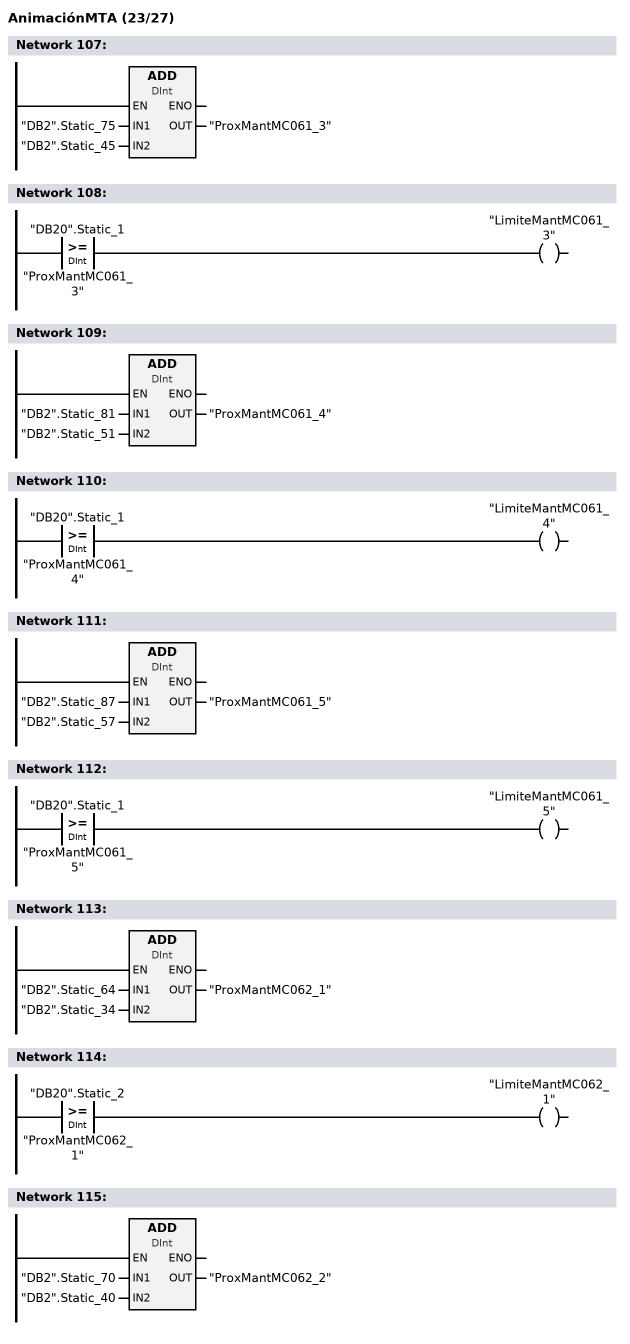
   RUNG wire#powerrail
      { S7_Templates := "SrcType := DInt"; S7_GenerateENO := "TRUE" } Add(in1 := "DB2".Static_75, in2 := "DB2".Static_45, out => "ProxMantMC061_3")
   END_RUNG
   // the same network as SCL:
   "ProxMantMC061_3" := "DB2".Static_75 + "DB2".Static_45;
END_REGION

REGION Network 108
   RUNG wire#powerrail
      { S7_Templates := "SrcType := DInt" } GE_Contact(in1 := "DB20".Static_1, in2 := "ProxMantMC061_3")
      Coil( "LimiteMantMC061_3" )
   END_RUNG
   // the same network as SCL:
   "LimiteMantMC061_3" := "DB20".Static_1 >= "ProxMantMC061_3";
END_REGION

REGION Network 109
   RUNG wire#powerrail
      { S7_Templates := "SrcType := DInt"; S7_GenerateENO := "TRUE" } Add(in1 := "DB2".Static_81, in2 := "DB2".Static_51, out => "ProxMantMC061_4")
   END_RUNG
   // the same network as SCL:
   "ProxMantMC061_4" := "DB2".Static_81 + "DB2".Static_51;
END_REGION

REGION Network 110
   RUNG wire#powerrail
      { S7_Templates := "SrcType := DInt" } GE_Contact(in1 := "DB20".Static_1, in2 := "ProxMantMC061_4")
      Coil( "LimiteMantMC061_4" )
   END_RUNG
   // the same network as SCL:
   "LimiteMantMC061_4" := "DB20".Static_1 >= "ProxMantMC061_4";
END_REGION

REGION Network 111
   RUNG wire#powerrail
      { S7_Templates := "SrcType := DInt"; S7_GenerateENO := "TRUE" } Add(in1 := "DB2".Static_87, in2 := "DB2".Static_57, out => "ProxMantMC061_5")
   END_RUNG
   // the same network as SCL:
   "ProxMantMC061_5" := "DB2".Static_87 + "DB2".Static_57;
END_REGION

REGION Network 112
   RUNG wire#powerrail
      { S7_Templates := "SrcType := DInt" } GE_Contact(in1 := "DB20".Static_1, in2 := "ProxMantMC061_5")
      Coil( "LimiteMantMC061_5" )
   END_RUNG
   // the same network as SCL:
   "LimiteMantMC061_5" := "DB20".Static_1 >= "ProxMantMC061_5";
END_REGION

REGION Network 113
   RUNG wire#powerrail
      { S7_Templates := "SrcType := DInt"; S7_GenerateENO := "TRUE" } Add(in1 := "DB2".Static_64, in2 := "DB2".Static_34, out => "ProxMantMC062_1")
   END_RUNG
   // the same network as SCL:
   "ProxMantMC062_1" := "DB2".Static_64 + "DB2".Static_34;
END_REGION

REGION Network 114
   RUNG wire#powerrail
      { S7_Templates := "SrcType := DInt" } GE_Contact(in1 := "DB20".Static_2, in2 := "ProxMantMC062_1")
      Coil( "LimiteMantMC062_1" )
   END_RUNG
   // the same network as SCL:
   "LimiteMantMC062_1" := "DB20".Static_2 >= "ProxMantMC062_1";
END_REGION

REGION Network 115
   RUNG wire#powerrail
      { S7_Templates := "SrcType := DInt"; S7_GenerateENO := "TRUE" } Add(in1 := "DB2".Static_70, in2 := "DB2".Static_40, out => "ProxMantMC062_2")
   END_RUNG
   // the same network as SCL:
   "ProxMantMC062_2" := "DB2".Static_70 + "DB2".Static_40;
END_REGION

REGION Network 116
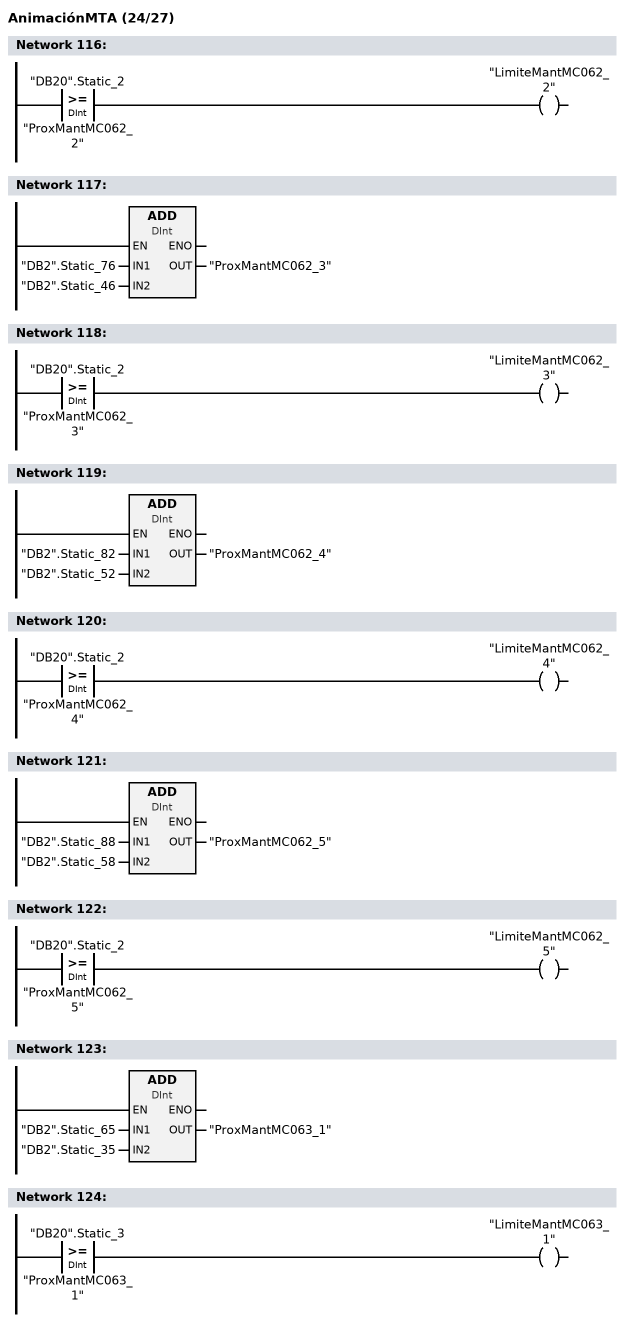
   RUNG wire#powerrail
      { S7_Templates := "SrcType := DInt" } GE_Contact(in1 := "DB20".Static_2, in2 := "ProxMantMC062_2")
      Coil( "LimiteMantMC062_2" )
   END_RUNG
   // the same network as SCL:
   "LimiteMantMC062_2" := "DB20".Static_2 >= "ProxMantMC062_2";
END_REGION

REGION Network 117
   RUNG wire#powerrail
      { S7_Templates := "SrcType := DInt"; S7_GenerateENO := "TRUE" } Add(in1 := "DB2".Static_76, in2 := "DB2".Static_46, out => "ProxMantMC062_3")
   END_RUNG
   // the same network as SCL:
   "ProxMantMC062_3" := "DB2".Static_76 + "DB2".Static_46;
END_REGION

REGION Network 118
   RUNG wire#powerrail
      { S7_Templates := "SrcType := DInt" } GE_Contact(in1 := "DB20".Static_2, in2 := "ProxMantMC062_3")
      Coil( "LimiteMantMC062_3" )
   END_RUNG
   // the same network as SCL:
   "LimiteMantMC062_3" := "DB20".Static_2 >= "ProxMantMC062_3";
END_REGION

REGION Network 119
   RUNG wire#powerrail
      { S7_Templates := "SrcType := DInt"; S7_GenerateENO := "TRUE" } Add(in1 := "DB2".Static_82, in2 := "DB2".Static_52, out => "ProxMantMC062_4")
   END_RUNG
   // the same network as SCL:
   "ProxMantMC062_4" := "DB2".Static_82 + "DB2".Static_52;
END_REGION

REGION Network 120
   RUNG wire#powerrail
      { S7_Templates := "SrcType := DInt" } GE_Contact(in1 := "DB20".Static_2, in2 := "ProxMantMC062_4")
      Coil( "LimiteMantMC062_4" )
   END_RUNG
   // the same network as SCL:
   "LimiteMantMC062_4" := "DB20".Static_2 >= "ProxMantMC062_4";
END_REGION

REGION Network 121
   RUNG wire#powerrail
      { S7_Templates := "SrcType := DInt"; S7_GenerateENO := "TRUE" } Add(in1 := "DB2".Static_88, in2 := "DB2".Static_58, out => "ProxMantMC062_5")
   END_RUNG
   // the same network as SCL:
   "ProxMantMC062_5" := "DB2".Static_88 + "DB2".Static_58;
END_REGION

REGION Network 122
   RUNG wire#powerrail
      { S7_Templates := "SrcType := DInt" } GE_Contact(in1 := "DB20".Static_2, in2 := "ProxMantMC062_5")
      Coil( "LimiteMantMC062_5" )
   END_RUNG
   // the same network as SCL:
   "LimiteMantMC062_5" := "DB20".Static_2 >= "ProxMantMC062_5";
END_REGION

REGION Network 123
   RUNG wire#powerrail
      { S7_Templates := "SrcType := DInt"; S7_GenerateENO := "TRUE" } Add(in1 := "DB2".Static_65, in2 := "DB2".Static_35, out => "ProxMantMC063_1")
   END_RUNG
   // the same network as SCL:
   "ProxMantMC063_1" := "DB2".Static_65 + "DB2".Static_35;
END_REGION

REGION Network 124
   RUNG wire#powerrail
      { S7_Templates := "SrcType := DInt" } GE_Contact(in1 := "DB20".Static_3, in2 := "ProxMantMC063_1")
      Coil( "LimiteMantMC063_1" )
   END_RUNG
   // the same network as SCL:
   "LimiteMantMC063_1" := "DB20".Static_3 >= "ProxMantMC063_1";
END_REGION

REGION Network 125
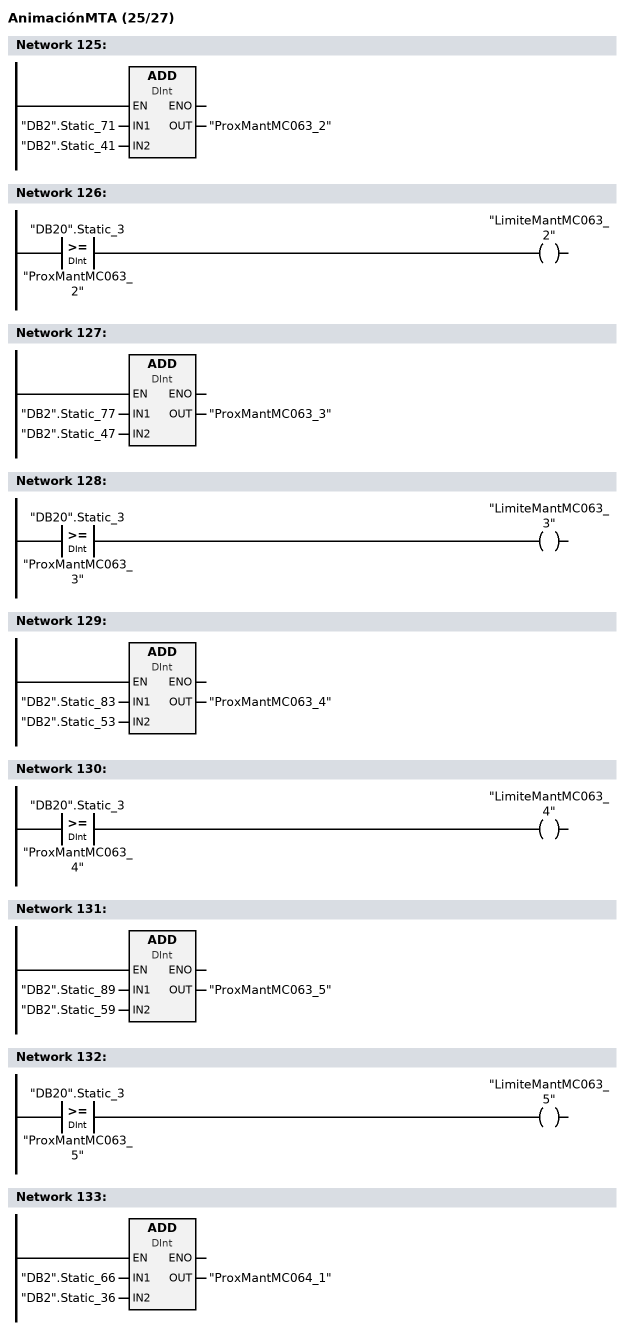
   RUNG wire#powerrail
      { S7_Templates := "SrcType := DInt"; S7_GenerateENO := "TRUE" } Add(in1 := "DB2".Static_71, in2 := "DB2".Static_41, out => "ProxMantMC063_2")
   END_RUNG
   // the same network as SCL:
   "ProxMantMC063_2" := "DB2".Static_71 + "DB2".Static_41;
END_REGION

REGION Network 126
   RUNG wire#powerrail
      { S7_Templates := "SrcType := DInt" } GE_Contact(in1 := "DB20".Static_3, in2 := "ProxMantMC063_2")
      Coil( "LimiteMantMC063_2" )
   END_RUNG
   // the same network as SCL:
   "LimiteMantMC063_2" := "DB20".Static_3 >= "ProxMantMC063_2";
END_REGION

REGION Network 127
   RUNG wire#powerrail
      { S7_Templates := "SrcType := DInt"; S7_GenerateENO := "TRUE" } Add(in1 := "DB2".Static_77, in2 := "DB2".Static_47, out => "ProxMantMC063_3")
   END_RUNG
   // the same network as SCL:
   "ProxMantMC063_3" := "DB2".Static_77 + "DB2".Static_47;
END_REGION

REGION Network 128
   RUNG wire#powerrail
      { S7_Templates := "SrcType := DInt" } GE_Contact(in1 := "DB20".Static_3, in2 := "ProxMantMC063_3")
      Coil( "LimiteMantMC063_3" )
   END_RUNG
   // the same network as SCL:
   "LimiteMantMC063_3" := "DB20".Static_3 >= "ProxMantMC063_3";
END_REGION

REGION Network 129
   RUNG wire#powerrail
      { S7_Templates := "SrcType := DInt"; S7_GenerateENO := "TRUE" } Add(in1 := "DB2".Static_83, in2 := "DB2".Static_53, out => "ProxMantMC063_4")
   END_RUNG
   // the same network as SCL:
   "ProxMantMC063_4" := "DB2".Static_83 + "DB2".Static_53;
END_REGION

REGION Network 130
   RUNG wire#powerrail
      { S7_Templates := "SrcType := DInt" } GE_Contact(in1 := "DB20".Static_3, in2 := "ProxMantMC063_4")
      Coil( "LimiteMantMC063_4" )
   END_RUNG
   // the same network as SCL:
   "LimiteMantMC063_4" := "DB20".Static_3 >= "ProxMantMC063_4";
END_REGION

REGION Network 131
   RUNG wire#powerrail
      { S7_Templates := "SrcType := DInt"; S7_GenerateENO := "TRUE" } Add(in1 := "DB2".Static_89, in2 := "DB2".Static_59, out => "ProxMantMC063_5")
   END_RUNG
   // the same network as SCL:
   "ProxMantMC063_5" := "DB2".Static_89 + "DB2".Static_59;
END_REGION

REGION Network 132
   RUNG wire#powerrail
      { S7_Templates := "SrcType := DInt" } GE_Contact(in1 := "DB20".Static_3, in2 := "ProxMantMC063_5")
      Coil( "LimiteMantMC063_5" )
   END_RUNG
   // the same network as SCL:
   "LimiteMantMC063_5" := "DB20".Static_3 >= "ProxMantMC063_5";
END_REGION

REGION Network 133
   RUNG wire#powerrail
      { S7_Templates := "SrcType := DInt"; S7_GenerateENO := "TRUE" } Add(in1 := "DB2".Static_66, in2 := "DB2".Static_36, out => "ProxMantMC064_1")
   END_RUNG
   // the same network as SCL:
   "ProxMantMC064_1" := "DB2".Static_66 + "DB2".Static_36;
END_REGION

REGION Network 134
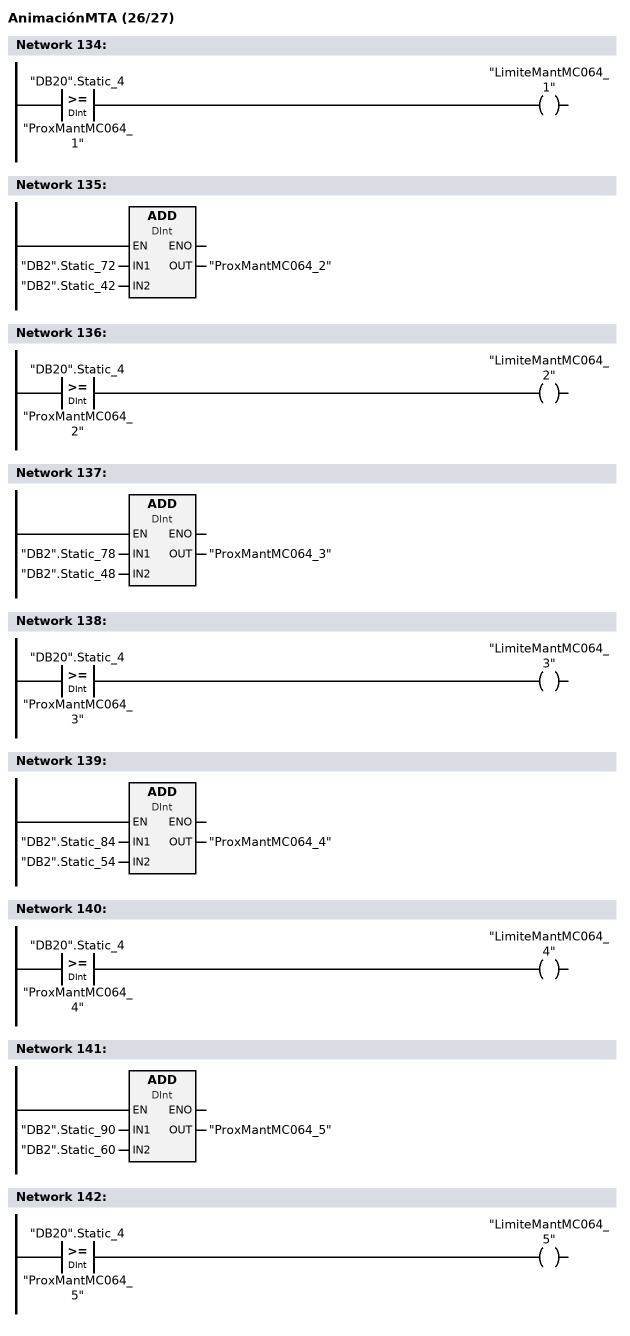
   RUNG wire#powerrail
      { S7_Templates := "SrcType := DInt" } GE_Contact(in1 := "DB20".Static_4, in2 := "ProxMantMC064_1")
      Coil( "LimiteMantMC064_1" )
   END_RUNG
   // the same network as SCL:
   "LimiteMantMC064_1" := "DB20".Static_4 >= "ProxMantMC064_1";
END_REGION

REGION Network 135
   RUNG wire#powerrail
      { S7_Templates := "SrcType := DInt"; S7_GenerateENO := "TRUE" } Add(in1 := "DB2".Static_72, in2 := "DB2".Static_42, out => "ProxMantMC064_2")
   END_RUNG
   // the same network as SCL:
   "ProxMantMC064_2" := "DB2".Static_72 + "DB2".Static_42;
END_REGION

REGION Network 136
   RUNG wire#powerrail
      { S7_Templates := "SrcType := DInt" } GE_Contact(in1 := "DB20".Static_4, in2 := "ProxMantMC064_2")
      Coil( "LimiteMantMC064_2" )
   END_RUNG
   // the same network as SCL:
   "LimiteMantMC064_2" := "DB20".Static_4 >= "ProxMantMC064_2";
END_REGION

REGION Network 137
   RUNG wire#powerrail
      { S7_Templates := "SrcType := DInt"; S7_GenerateENO := "TRUE" } Add(in1 := "DB2".Static_78, in2 := "DB2".Static_48, out => "ProxMantMC064_3")
   END_RUNG
   // the same network as SCL:
   "ProxMantMC064_3" := "DB2".Static_78 + "DB2".Static_48;
END_REGION

REGION Network 138
   RUNG wire#powerrail
      { S7_Templates := "SrcType := DInt" } GE_Contact(in1 := "DB20".Static_4, in2 := "ProxMantMC064_3")
      Coil( "LimiteMantMC064_3" )
   END_RUNG
   // the same network as SCL:
   "LimiteMantMC064_3" := "DB20".Static_4 >= "ProxMantMC064_3";
END_REGION

REGION Network 139
   RUNG wire#powerrail
      { S7_Templates := "SrcType := DInt"; S7_GenerateENO := "TRUE" } Add(in1 := "DB2".Static_84, in2 := "DB2".Static_54, out => "ProxMantMC064_4")
   END_RUNG
   // the same network as SCL:
   "ProxMantMC064_4" := "DB2".Static_84 + "DB2".Static_54;
END_REGION

REGION Network 140
   RUNG wire#powerrail
      { S7_Templates := "SrcType := DInt" } GE_Contact(in1 := "DB20".Static_4, in2 := "ProxMantMC064_4")
      Coil( "LimiteMantMC064_4" )
   END_RUNG
   // the same network as SCL:
   "LimiteMantMC064_4" := "DB20".Static_4 >= "ProxMantMC064_4";
END_REGION

REGION Network 141
   RUNG wire#powerrail
      { S7_Templates := "SrcType := DInt"; S7_GenerateENO := "TRUE" } Add(in1 := "DB2".Static_90, in2 := "DB2".Static_60, out => "ProxMantMC064_5")
   END_RUNG
   // the same network as SCL:
   "ProxMantMC064_5" := "DB2".Static_90 + "DB2".Static_60;
END_REGION

REGION Network 142
   RUNG wire#powerrail
      { S7_Templates := "SrcType := DInt" } GE_Contact(in1 := "DB20".Static_4, in2 := "ProxMantMC064_5")
      Coil( "LimiteMantMC064_5" )
   END_RUNG
   // the same network as SCL:
   "LimiteMantMC064_5" := "DB20".Static_4 >= "ProxMantMC064_5";
END_REGION

REGION Network 143
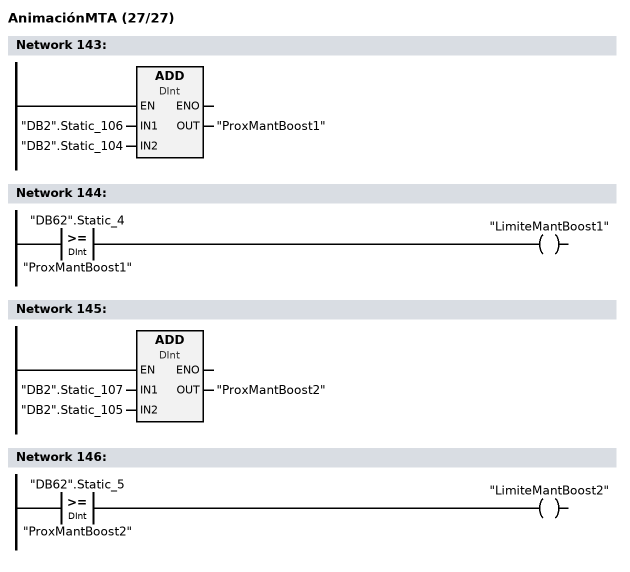
   RUNG wire#powerrail
      { S7_Templates := "SrcType := DInt"; S7_GenerateENO := "TRUE" } Add(in1 := "DB2".Static_106, in2 := "DB2".Static_104, out => "ProxMantBoost1")
   END_RUNG
   // the same network as SCL:
   "ProxMantBoost1" := "DB2".Static_106 + "DB2".Static_104;
END_REGION

REGION Network 144
   RUNG wire#powerrail
      { S7_Templates := "SrcType := DInt" } GE_Contact(in1 := "DB62".Static_4, in2 := "ProxMantBoost1")
      Coil( "LimiteMantBoost1" )
   END_RUNG
   // the same network as SCL:
   "LimiteMantBoost1" := "DB62".Static_4 >= "ProxMantBoost1";
END_REGION

REGION Network 145
   RUNG wire#powerrail
      { S7_Templates := "SrcType := DInt"; S7_GenerateENO := "TRUE" } Add(in1 := "DB2".Static_107, in2 := "DB2".Static_105, out => "ProxMantBoost2")
   END_RUNG
   // the same network as SCL:
   "ProxMantBoost2" := "DB2".Static_107 + "DB2".Static_105;
END_REGION

REGION Network 146
   RUNG wire#powerrail
      { S7_Templates := "SrcType := DInt" } GE_Contact(in1 := "DB62".Static_5, in2 := "ProxMantBoost2")
      Coil( "LimiteMantBoost2" )
   END_RUNG
   // the same network as SCL:
   "LimiteMantBoost2" := "DB62".Static_5 >= "ProxMantBoost2";
END_REGION
END_FUNCTION

FUNCTION "Motores-PanelMTA" : Void   // FC3, LAD
{ S7_Optimized_Access := 'FALSE' }
VERSION : 0.1
BEGIN

REGION Network 1
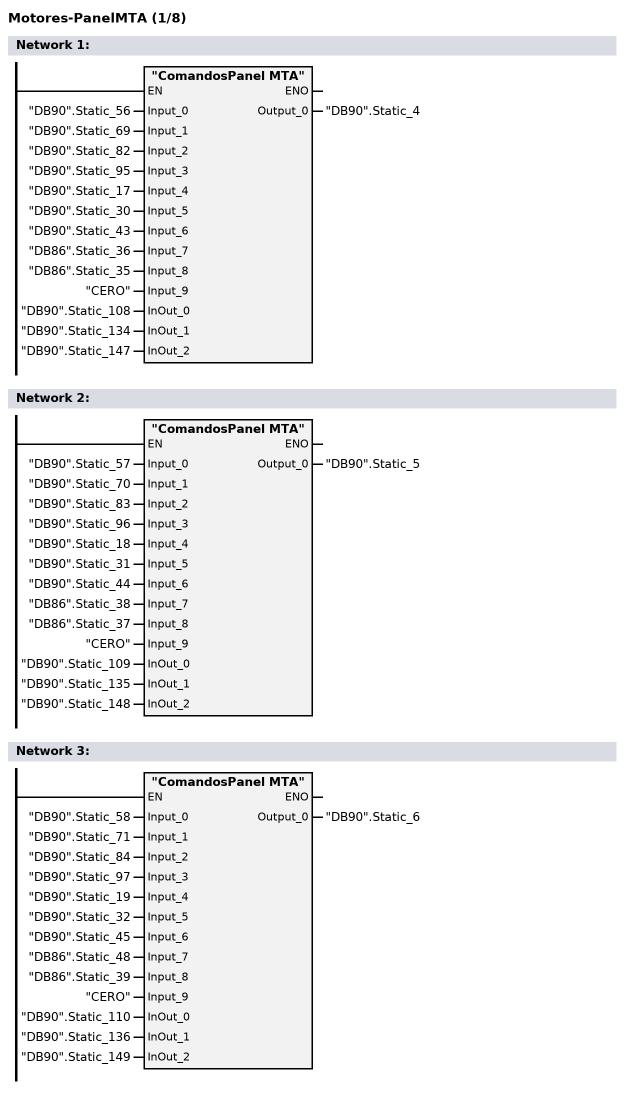
   RUNG wire#powerrail
      "ComandosPanel MTA"(Input_0 := "DB90".Static_56, Input_1 := "DB90".Static_69, Input_2 := "DB90".Static_82, Input_3 := "DB90".Static_95, Input_4 := "DB90".Static_17, Input_5 := "DB90".Static_30, Input_6 := "DB90".Static_43, Input_7 := "DB86".Static_36, Input_8 := "DB86".Static_35, Input_9 := "CERO", Output_0 => "DB90".Static_4, InOut_0 := "DB90".Static_108, InOut_1 := "DB90".Static_134, InOut_2 := "DB90".Static_147)
   END_RUNG
   // the same network as SCL:
   "ComandosPanel MTA"(Input_0 := "DB90".Static_56,
                       Input_1 := "DB90".Static_69,
                       Input_2 := "DB90".Static_82,
                       Input_3 := "DB90".Static_95,
                       Input_4 := "DB90".Static_17,
                       Input_5 := "DB90".Static_30,
                       Input_6 := "DB90".Static_43,
                       Input_7 := "DB86".Static_36,
                       Input_8 := "DB86".Static_35,
                       Input_9 := "CERO",
                       InOut_0 := "DB90".Static_108,
                       InOut_1 := "DB90".Static_134,
                       InOut_2 := "DB90".Static_147,
                       Output_0 => "DB90".Static_4);
END_REGION

REGION Network 2
   RUNG wire#powerrail
      "ComandosPanel MTA"(Input_0 := "DB90".Static_57, Input_1 := "DB90".Static_70, Input_2 := "DB90".Static_83, Input_3 := "DB90".Static_96, Input_4 := "DB90".Static_18, Input_5 := "DB90".Static_31, Input_6 := "DB90".Static_44, Input_7 := "DB86".Static_38, Input_8 := "DB86".Static_37, Input_9 := "CERO", Output_0 => "DB90".Static_5, InOut_0 := "DB90".Static_109, InOut_1 := "DB90".Static_135, InOut_2 := "DB90".Static_148)
   END_RUNG
   // the same network as SCL:
   "ComandosPanel MTA"(Input_0 := "DB90".Static_57,
                       Input_1 := "DB90".Static_70,
                       Input_2 := "DB90".Static_83,
                       Input_3 := "DB90".Static_96,
                       Input_4 := "DB90".Static_18,
                       Input_5 := "DB90".Static_31,
                       Input_6 := "DB90".Static_44,
                       Input_7 := "DB86".Static_38,
                       Input_8 := "DB86".Static_37,
                       Input_9 := "CERO",
                       InOut_0 := "DB90".Static_109,
                       InOut_1 := "DB90".Static_135,
                       InOut_2 := "DB90".Static_148,
                       Output_0 => "DB90".Static_5);
END_REGION

REGION Network 3
   RUNG wire#powerrail
      "ComandosPanel MTA"(Input_0 := "DB90".Static_58, Input_1 := "DB90".Static_71, Input_2 := "DB90".Static_84, Input_3 := "DB90".Static_97, Input_4 := "DB90".Static_19, Input_5 := "DB90".Static_32, Input_6 := "DB90".Static_45, Input_7 := "DB86".Static_48, Input_8 := "DB86".Static_39, Input_9 := "CERO", Output_0 => "DB90".Static_6, InOut_0 := "DB90".Static_110, InOut_1 := "DB90".Static_136, InOut_2 := "DB90".Static_149)
   END_RUNG
   // the same network as SCL:
   "ComandosPanel MTA"(Input_0 := "DB90".Static_58,
                       Input_1 := "DB90".Static_71,
                       Input_2 := "DB90".Static_84,
                       Input_3 := "DB90".Static_97,
                       Input_4 := "DB90".Static_19,
                       Input_5 := "DB90".Static_32,
                       Input_6 := "DB90".Static_45,
                       Input_7 := "DB86".Static_48,
                       Input_8 := "DB86".Static_39,
                       Input_9 := "CERO",
                       InOut_0 := "DB90".Static_110,
                       InOut_1 := "DB90".Static_136,
                       InOut_2 := "DB90".Static_149,
                       Output_0 => "DB90".Static_6);
END_REGION

REGION Network 4
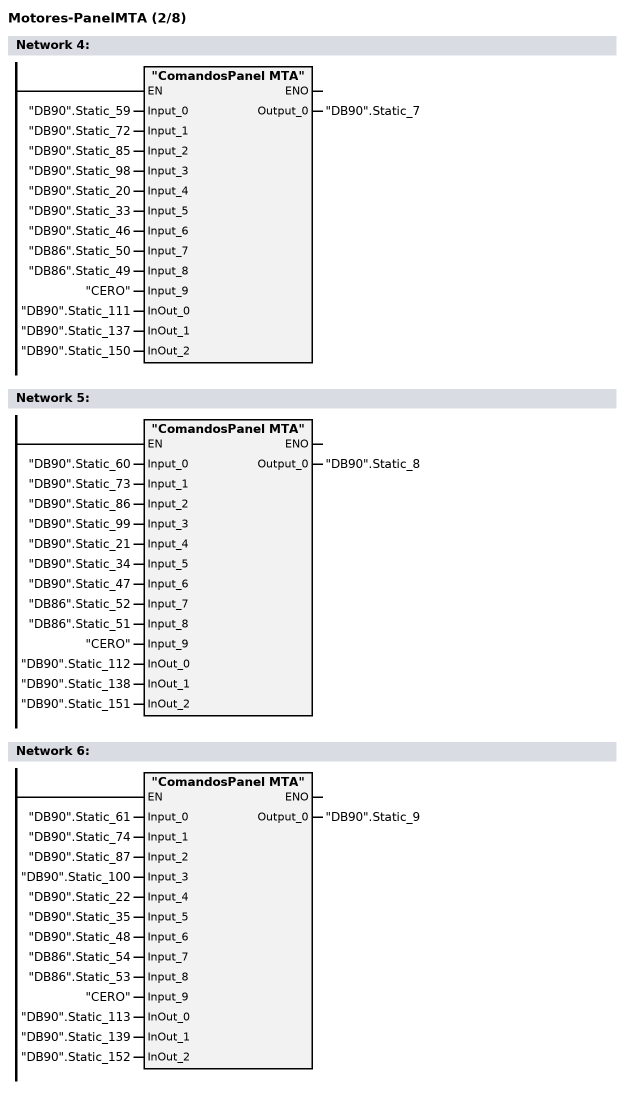
   RUNG wire#powerrail
      "ComandosPanel MTA"(Input_0 := "DB90".Static_59, Input_1 := "DB90".Static_72, Input_2 := "DB90".Static_85, Input_3 := "DB90".Static_98, Input_4 := "DB90".Static_20, Input_5 := "DB90".Static_33, Input_6 := "DB90".Static_46, Input_7 := "DB86".Static_50, Input_8 := "DB86".Static_49, Input_9 := "CERO", Output_0 => "DB90".Static_7, InOut_0 := "DB90".Static_111, InOut_1 := "DB90".Static_137, InOut_2 := "DB90".Static_150)
   END_RUNG
   // the same network as SCL:
   "ComandosPanel MTA"(Input_0 := "DB90".Static_59,
                       Input_1 := "DB90".Static_72,
                       Input_2 := "DB90".Static_85,
                       Input_3 := "DB90".Static_98,
                       Input_4 := "DB90".Static_20,
                       Input_5 := "DB90".Static_33,
                       Input_6 := "DB90".Static_46,
                       Input_7 := "DB86".Static_50,
                       Input_8 := "DB86".Static_49,
                       Input_9 := "CERO",
                       InOut_0 := "DB90".Static_111,
                       InOut_1 := "DB90".Static_137,
                       InOut_2 := "DB90".Static_150,
                       Output_0 => "DB90".Static_7);
END_REGION

REGION Network 5
   RUNG wire#powerrail
      "ComandosPanel MTA"(Input_0 := "DB90".Static_60, Input_1 := "DB90".Static_73, Input_2 := "DB90".Static_86, Input_3 := "DB90".Static_99, Input_4 := "DB90".Static_21, Input_5 := "DB90".Static_34, Input_6 := "DB90".Static_47, Input_7 := "DB86".Static_52, Input_8 := "DB86".Static_51, Input_9 := "CERO", Output_0 => "DB90".Static_8, InOut_0 := "DB90".Static_112, InOut_1 := "DB90".Static_138, InOut_2 := "DB90".Static_151)
   END_RUNG
   // the same network as SCL:
   "ComandosPanel MTA"(Input_0 := "DB90".Static_60,
                       Input_1 := "DB90".Static_73,
                       Input_2 := "DB90".Static_86,
                       Input_3 := "DB90".Static_99,
                       Input_4 := "DB90".Static_21,
                       Input_5 := "DB90".Static_34,
                       Input_6 := "DB90".Static_47,
                       Input_7 := "DB86".Static_52,
                       Input_8 := "DB86".Static_51,
                       Input_9 := "CERO",
                       InOut_0 := "DB90".Static_112,
                       InOut_1 := "DB90".Static_138,
                       InOut_2 := "DB90".Static_151,
                       Output_0 => "DB90".Static_8);
END_REGION

REGION Network 6
   RUNG wire#powerrail
      "ComandosPanel MTA"(Input_0 := "DB90".Static_61, Input_1 := "DB90".Static_74, Input_2 := "DB90".Static_87, Input_3 := "DB90".Static_100, Input_4 := "DB90".Static_22, Input_5 := "DB90".Static_35, Input_6 := "DB90".Static_48, Input_7 := "DB86".Static_54, Input_8 := "DB86".Static_53, Input_9 := "CERO", Output_0 => "DB90".Static_9, InOut_0 := "DB90".Static_113, InOut_1 := "DB90".Static_139, InOut_2 := "DB90".Static_152)
   END_RUNG
   // the same network as SCL:
   "ComandosPanel MTA"(Input_0 := "DB90".Static_61,
                       Input_1 := "DB90".Static_74,
                       Input_2 := "DB90".Static_87,
                       Input_3 := "DB90".Static_100,
                       Input_4 := "DB90".Static_22,
                       Input_5 := "DB90".Static_35,
                       Input_6 := "DB90".Static_48,
                       Input_7 := "DB86".Static_54,
                       Input_8 := "DB86".Static_53,
                       Input_9 := "CERO",
                       InOut_0 := "DB90".Static_113,
                       InOut_1 := "DB90".Static_139,
                       InOut_2 := "DB90".Static_152,
                       Output_0 => "DB90".Static_9);
END_REGION

REGION Network 7
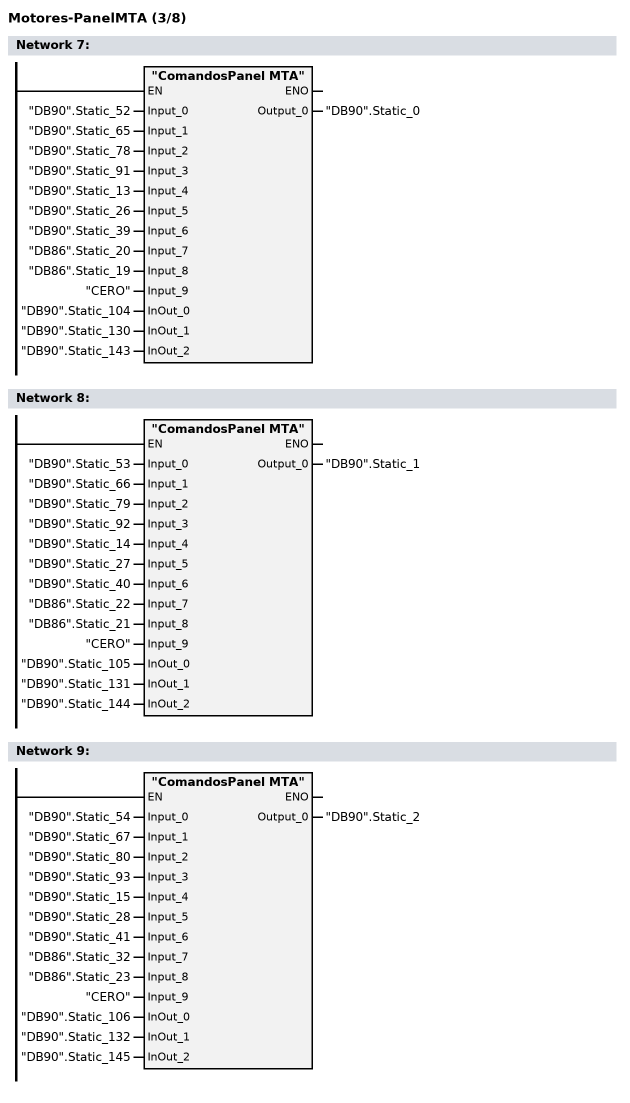
   RUNG wire#powerrail
      "ComandosPanel MTA"(Input_0 := "DB90".Static_52, Input_1 := "DB90".Static_65, Input_2 := "DB90".Static_78, Input_3 := "DB90".Static_91, Input_4 := "DB90".Static_13, Input_5 := "DB90".Static_26, Input_6 := "DB90".Static_39, Input_7 := "DB86".Static_20, Input_8 := "DB86".Static_19, Input_9 := "CERO", Output_0 => "DB90".Static_0, InOut_0 := "DB90".Static_104, InOut_1 := "DB90".Static_130, InOut_2 := "DB90".Static_143)
   END_RUNG
   // the same network as SCL:
   "ComandosPanel MTA"(Input_0 := "DB90".Static_52,
                       Input_1 := "DB90".Static_65,
                       Input_2 := "DB90".Static_78,
                       Input_3 := "DB90".Static_91,
                       Input_4 := "DB90".Static_13,
                       Input_5 := "DB90".Static_26,
                       Input_6 := "DB90".Static_39,
                       Input_7 := "DB86".Static_20,
                       Input_8 := "DB86".Static_19,
                       Input_9 := "CERO",
                       InOut_0 := "DB90".Static_104,
                       InOut_1 := "DB90".Static_130,
                       InOut_2 := "DB90".Static_143,
                       Output_0 => "DB90".Static_0);
END_REGION

REGION Network 8
   RUNG wire#powerrail
      "ComandosPanel MTA"(Input_0 := "DB90".Static_53, Input_1 := "DB90".Static_66, Input_2 := "DB90".Static_79, Input_3 := "DB90".Static_92, Input_4 := "DB90".Static_14, Input_5 := "DB90".Static_27, Input_6 := "DB90".Static_40, Input_7 := "DB86".Static_22, Input_8 := "DB86".Static_21, Input_9 := "CERO", Output_0 => "DB90".Static_1, InOut_0 := "DB90".Static_105, InOut_1 := "DB90".Static_131, InOut_2 := "DB90".Static_144)
   END_RUNG
   // the same network as SCL:
   "ComandosPanel MTA"(Input_0 := "DB90".Static_53,
                       Input_1 := "DB90".Static_66,
                       Input_2 := "DB90".Static_79,
                       Input_3 := "DB90".Static_92,
                       Input_4 := "DB90".Static_14,
                       Input_5 := "DB90".Static_27,
                       Input_6 := "DB90".Static_40,
                       Input_7 := "DB86".Static_22,
                       Input_8 := "DB86".Static_21,
                       Input_9 := "CERO",
                       InOut_0 := "DB90".Static_105,
                       InOut_1 := "DB90".Static_131,
                       InOut_2 := "DB90".Static_144,
                       Output_0 => "DB90".Static_1);
END_REGION

REGION Network 9
   RUNG wire#powerrail
      "ComandosPanel MTA"(Input_0 := "DB90".Static_54, Input_1 := "DB90".Static_67, Input_2 := "DB90".Static_80, Input_3 := "DB90".Static_93, Input_4 := "DB90".Static_15, Input_5 := "DB90".Static_28, Input_6 := "DB90".Static_41, Input_7 := "DB86".Static_32, Input_8 := "DB86".Static_23, Input_9 := "CERO", Output_0 => "DB90".Static_2, InOut_0 := "DB90".Static_106, InOut_1 := "DB90".Static_132, InOut_2 := "DB90".Static_145)
   END_RUNG
   // the same network as SCL:
   "ComandosPanel MTA"(Input_0 := "DB90".Static_54,
                       Input_1 := "DB90".Static_67,
                       Input_2 := "DB90".Static_80,
                       Input_3 := "DB90".Static_93,
                       Input_4 := "DB90".Static_15,
                       Input_5 := "DB90".Static_28,
                       Input_6 := "DB90".Static_41,
                       Input_7 := "DB86".Static_32,
                       Input_8 := "DB86".Static_23,
                       Input_9 := "CERO",
                       InOut_0 := "DB90".Static_106,
                       InOut_1 := "DB90".Static_132,
                       InOut_2 := "DB90".Static_145,
                       Output_0 => "DB90".Static_2);
END_REGION

REGION Network 10
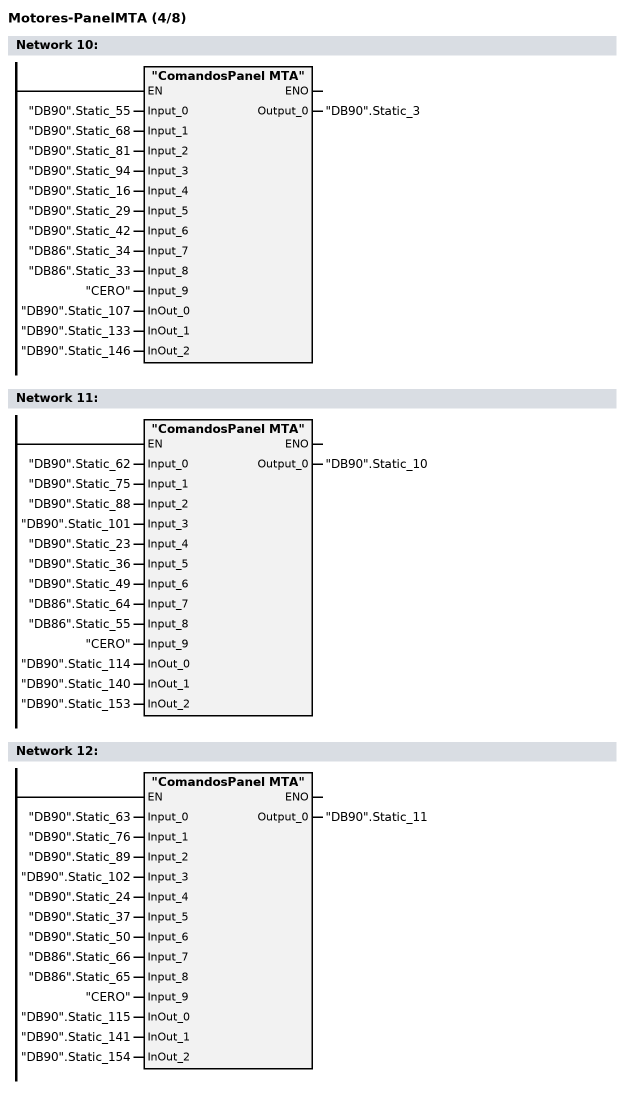
   RUNG wire#powerrail
      "ComandosPanel MTA"(Input_0 := "DB90".Static_55, Input_1 := "DB90".Static_68, Input_2 := "DB90".Static_81, Input_3 := "DB90".Static_94, Input_4 := "DB90".Static_16, Input_5 := "DB90".Static_29, Input_6 := "DB90".Static_42, Input_7 := "DB86".Static_34, Input_8 := "DB86".Static_33, Input_9 := "CERO", Output_0 => "DB90".Static_3, InOut_0 := "DB90".Static_107, InOut_1 := "DB90".Static_133, InOut_2 := "DB90".Static_146)
   END_RUNG
   // the same network as SCL:
   "ComandosPanel MTA"(Input_0 := "DB90".Static_55,
                       Input_1 := "DB90".Static_68,
                       Input_2 := "DB90".Static_81,
                       Input_3 := "DB90".Static_94,
                       Input_4 := "DB90".Static_16,
                       Input_5 := "DB90".Static_29,
                       Input_6 := "DB90".Static_42,
                       Input_7 := "DB86".Static_34,
                       Input_8 := "DB86".Static_33,
                       Input_9 := "CERO",
                       InOut_0 := "DB90".Static_107,
                       InOut_1 := "DB90".Static_133,
                       InOut_2 := "DB90".Static_146,
                       Output_0 => "DB90".Static_3);
END_REGION

REGION Network 11
   RUNG wire#powerrail
      "ComandosPanel MTA"(Input_0 := "DB90".Static_62, Input_1 := "DB90".Static_75, Input_2 := "DB90".Static_88, Input_3 := "DB90".Static_101, Input_4 := "DB90".Static_23, Input_5 := "DB90".Static_36, Input_6 := "DB90".Static_49, Input_7 := "DB86".Static_64, Input_8 := "DB86".Static_55, Input_9 := "CERO", Output_0 => "DB90".Static_10, InOut_0 := "DB90".Static_114, InOut_1 := "DB90".Static_140, InOut_2 := "DB90".Static_153)
   END_RUNG
   // the same network as SCL:
   "ComandosPanel MTA"(Input_0 := "DB90".Static_62,
                       Input_1 := "DB90".Static_75,
                       Input_2 := "DB90".Static_88,
                       Input_3 := "DB90".Static_101,
                       Input_4 := "DB90".Static_23,
                       Input_5 := "DB90".Static_36,
                       Input_6 := "DB90".Static_49,
                       Input_7 := "DB86".Static_64,
                       Input_8 := "DB86".Static_55,
                       Input_9 := "CERO",
                       InOut_0 := "DB90".Static_114,
                       InOut_1 := "DB90".Static_140,
                       InOut_2 := "DB90".Static_153,
                       Output_0 => "DB90".Static_10);
END_REGION

REGION Network 12
   RUNG wire#powerrail
      "ComandosPanel MTA"(Input_0 := "DB90".Static_63, Input_1 := "DB90".Static_76, Input_2 := "DB90".Static_89, Input_3 := "DB90".Static_102, Input_4 := "DB90".Static_24, Input_5 := "DB90".Static_37, Input_6 := "DB90".Static_50, Input_7 := "DB86".Static_66, Input_8 := "DB86".Static_65, Input_9 := "CERO", Output_0 => "DB90".Static_11, InOut_0 := "DB90".Static_115, InOut_1 := "DB90".Static_141, InOut_2 := "DB90".Static_154)
   END_RUNG
   // the same network as SCL:
   "ComandosPanel MTA"(Input_0 := "DB90".Static_63,
                       Input_1 := "DB90".Static_76,
                       Input_2 := "DB90".Static_89,
                       Input_3 := "DB90".Static_102,
                       Input_4 := "DB90".Static_24,
                       Input_5 := "DB90".Static_37,
                       Input_6 := "DB90".Static_50,
                       Input_7 := "DB86".Static_66,
                       Input_8 := "DB86".Static_65,
                       Input_9 := "CERO",
                       InOut_0 := "DB90".Static_115,
                       InOut_1 := "DB90".Static_141,
                       InOut_2 := "DB90".Static_154,
                       Output_0 => "DB90".Static_11);
END_REGION

REGION Network 13
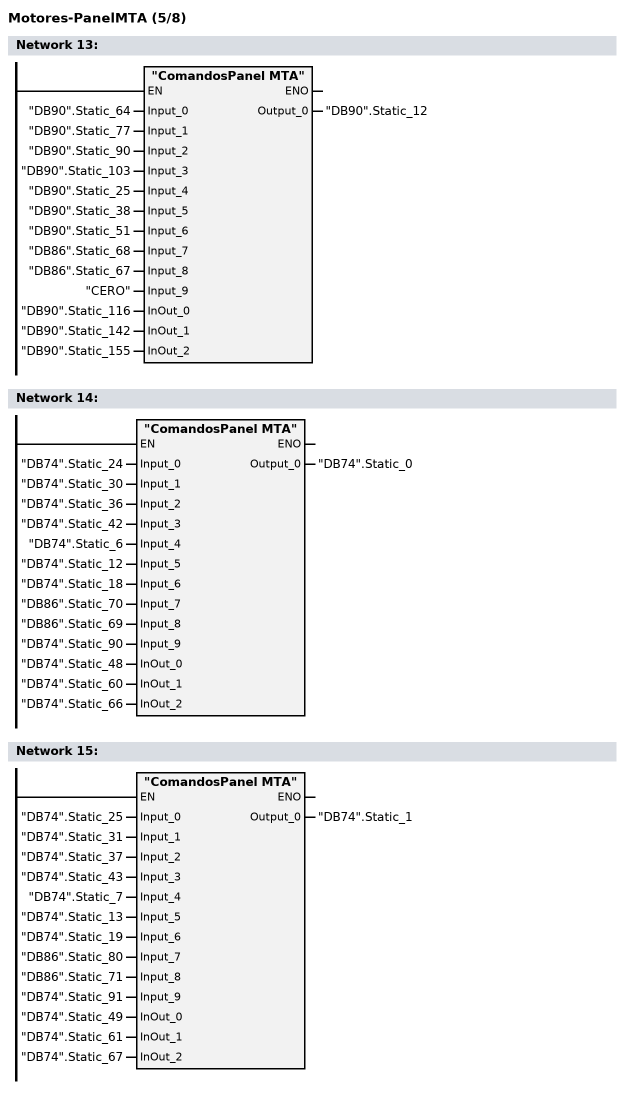
   RUNG wire#powerrail
      "ComandosPanel MTA"(Input_0 := "DB90".Static_64, Input_1 := "DB90".Static_77, Input_2 := "DB90".Static_90, Input_3 := "DB90".Static_103, Input_4 := "DB90".Static_25, Input_5 := "DB90".Static_38, Input_6 := "DB90".Static_51, Input_7 := "DB86".Static_68, Input_8 := "DB86".Static_67, Input_9 := "CERO", Output_0 => "DB90".Static_12, InOut_0 := "DB90".Static_116, InOut_1 := "DB90".Static_142, InOut_2 := "DB90".Static_155)
   END_RUNG
   // the same network as SCL:
   "ComandosPanel MTA"(Input_0 := "DB90".Static_64,
                       Input_1 := "DB90".Static_77,
                       Input_2 := "DB90".Static_90,
                       Input_3 := "DB90".Static_103,
                       Input_4 := "DB90".Static_25,
                       Input_5 := "DB90".Static_38,
                       Input_6 := "DB90".Static_51,
                       Input_7 := "DB86".Static_68,
                       Input_8 := "DB86".Static_67,
                       Input_9 := "CERO",
                       InOut_0 := "DB90".Static_116,
                       InOut_1 := "DB90".Static_142,
                       InOut_2 := "DB90".Static_155,
                       Output_0 => "DB90".Static_12);
END_REGION

REGION Network 14
   RUNG wire#powerrail
      "ComandosPanel MTA"(Input_0 := "DB74".Static_24, Input_1 := "DB74".Static_30, Input_2 := "DB74".Static_36, Input_3 := "DB74".Static_42, Input_4 := "DB74".Static_6, Input_5 := "DB74".Static_12, Input_6 := "DB74".Static_18, Input_7 := "DB86".Static_70, Input_8 := "DB86".Static_69, Input_9 := "DB74".Static_90, Output_0 => "DB74".Static_0, InOut_0 := "DB74".Static_48, InOut_1 := "DB74".Static_60, InOut_2 := "DB74".Static_66)
   END_RUNG
   // the same network as SCL:
   "ComandosPanel MTA"(Input_0 := "DB74".Static_24,
                       Input_1 := "DB74".Static_30,
                       Input_2 := "DB74".Static_36,
                       Input_3 := "DB74".Static_42,
                       Input_4 := "DB74".Static_6,
                       Input_5 := "DB74".Static_12,
                       Input_6 := "DB74".Static_18,
                       Input_7 := "DB86".Static_70,
                       Input_8 := "DB86".Static_69,
                       Input_9 := "DB74".Static_90,
                       InOut_0 := "DB74".Static_48,
                       InOut_1 := "DB74".Static_60,
                       InOut_2 := "DB74".Static_66,
                       Output_0 => "DB74".Static_0);
END_REGION

REGION Network 15
   RUNG wire#powerrail
      "ComandosPanel MTA"(Input_0 := "DB74".Static_25, Input_1 := "DB74".Static_31, Input_2 := "DB74".Static_37, Input_3 := "DB74".Static_43, Input_4 := "DB74".Static_7, Input_5 := "DB74".Static_13, Input_6 := "DB74".Static_19, Input_7 := "DB86".Static_80, Input_8 := "DB86".Static_71, Input_9 := "DB74".Static_91, Output_0 => "DB74".Static_1, InOut_0 := "DB74".Static_49, InOut_1 := "DB74".Static_61, InOut_2 := "DB74".Static_67)
   END_RUNG
   // the same network as SCL:
   "ComandosPanel MTA"(Input_0 := "DB74".Static_25,
                       Input_1 := "DB74".Static_31,
                       Input_2 := "DB74".Static_37,
                       Input_3 := "DB74".Static_43,
                       Input_4 := "DB74".Static_7,
                       Input_5 := "DB74".Static_13,
                       Input_6 := "DB74".Static_19,
                       Input_7 := "DB86".Static_80,
                       Input_8 := "DB86".Static_71,
                       Input_9 := "DB74".Static_91,
                       InOut_0 := "DB74".Static_49,
                       InOut_1 := "DB74".Static_61,
                       InOut_2 := "DB74".Static_67,
                       Output_0 => "DB74".Static_1);
END_REGION

REGION Network 16